   
   //M307EM1
   Z300_Conveyor_Conf[19].dLengthConveyor_cmm := 238000;
   Z300_Conveyor_Conf[19].dWidthConveyor_cmm := 450000;
   Z300_Conveyor_Conf[19].dPitchRoller := 25000;
   Z300_Conveyor_Conf[19].dSpaceRestartPlate_cmm := 200000;
   Z300_Conveyor_Conf[19].dMachineIndex := 19;
   Z300_Conveyor_Conf[19].dZoneConveyor := 1; //Z301
   Z300_Conveyor_Conf[19].dMotorNumber := 0; //Single motor
   Z300_Conveyor_Conf[19].dIndexMainSpeed := 0; //Auto speed
   Z300_Conveyor_Conf[19].xContinuousConveyor := 0;
   Z300_Conveyor_Conf[19].xWaitGlassForStop := 1;
   Z300_Conveyor_Conf[19].rAccH_ms2 := 1.2;
   Z300_Conveyor_Conf[19].rDecH_ms2 := 1.2;
   Z300_Conveyor_Conf[19].rAccH_s := 1.25; //acceleration time with max speed 90 m/min
   Z300_Conveyor_Conf[19].rDecH_s := 1.25; //acceleration time with max speed 90 m/min
   Z300_Conveyor_Conf[19].rAccL_ms2 := 0.7;
   Z300_Conveyor_Conf[19].rDecL_ms2 := 0.7;
   Z300_Conveyor_Conf[19].rAccL_s := 2.14; //acceleration time with max speed 90 m/min
   Z300_Conveyor_Conf[19].rDecL_s := 2.14; //acceleration time with max speed 90 m/min
   Z300_Conveyor_Conf[19].xSimulationMotor := TMP_xSimulationActive;
   Z300_Conveyor_Conf[19].xLocalCleaningAllow := 0;
   Z300_Conveyor_Conf[19].xOnlyOnePlateAtTheTime := 0;
   Z300_Conveyor_Conf[19].rgxAllowedDest := CONST_rgdDestMask[0] AND CONST_rgdDestMask[1] AND CONST_rgdDestMask[2] AND CONST_rgdDestMask[3] AND CONST_rgdDestMask[4] AND CONST_rgdDestMask[5] AND CONST_rgdDestMask[6];
   Z300_Conveyor_Conf[19].rgxAllowedCullet := CONST_rgdDestMask[24];
   Z300_Conveyor_Conf[19].rgxAllowedQuality := CONST_rgdDestMask[29] AND CONST_rgdDestMask[30] AND CONST_rgdDestMask[31];
   Z300_Conveyor[19].tmOFF_DriveEnable[0].PRE := 30000;
   Z300_Conveyor[19].tmON_FeedbackTimeout[0].PRE := 2500;
   Z300_Conveyor[19].tmON_FeedbackTimeout[1].PRE := 2500;
   Z300_Conveyor[19].tmON_DelayReadyToMove[0].PRE := 200;
   Z300_Conveyor[19].tmON_DelayReadyToMove[1].PRE := 200;
   Z300_Conveyor[19].tmON_FeedbackDriveReady[0].PRE := 1000;
   Z300_Conveyor[19].tmON_FeedbackDriveReady[1].PRE := 1000;
   
   //M307FM1
   Z300_Conveyor_Conf[20].dLengthConveyor_cmm := 238000;
   Z300_Conveyor_Conf[20].dWidthConveyor_cmm := 450000;
   Z300_Conveyor_Conf[20].dPitchRoller := 25000;
   Z300_Conveyor_Conf[20].dSpaceRestartPlate_cmm := 200000;
   Z300_Conveyor_Conf[20].dMachineIndex := 20;
   Z300_Conveyor_Conf[20].dZoneConveyor := 1; //Z301
   Z300_Conveyor_Conf[20].dMotorNumber := 0; //Single motor
   Z300_Conveyor_Conf[20].dIndexMainSpeed := 0; //Auto speed
   Z300_Conveyor_Conf[20].xContinuousConveyor := 0;
   Z300_Conveyor_Conf[20].xWaitGlassForStop := 1;
   Z300_Conveyor_Conf[20].rAccH_ms2 := 1.2;
   Z300_Conveyor_Conf[20].rDecH_ms2 := 1.2;
   Z300_Conveyor_Conf[20].rAccH_s := 1.25; //acceleration time with max speed 90 m/min
   Z300_Conveyor_Conf[20].rDecH_s := 1.25; //acceleration time with max speed 90 m/min
   Z300_Conveyor_Conf[20].rAccL_ms2 := 0.7;
   Z300_Conveyor_Conf[20].rDecL_ms2 := 0.7;
   Z300_Conveyor_Conf[20].rAccL_s := 2.14; //acceleration time with max speed 90 m/min
   Z300_Conveyor_Conf[20].rDecL_s := 2.14; //acceleration time with max speed 90 m/min
   Z300_Conveyor_Conf[20].xSimulationMotor := TMP_xSimulationActive;
   Z300_Conveyor_Conf[20].xLocalCleaningAllow := 0;
   Z300_Conveyor_Conf[20].xOnlyOnePlateAtTheTime := 0;
   Z300_Conveyor_Conf[20].rgxAllowedDest := CONST_rgdDestMask[0] AND CONST_rgdDestMask[1] AND CONST_rgdDestMask[2] AND CONST_rgdDestMask[3] AND CONST_rgdDestMask[4] AND CONST_rgdDestMask[5] AND CONST_rgdDestMask[6];
   Z300_Conveyor_Conf[20].rgxAllowedCullet := CONST_rgdDestMask[24];
   Z300_Conveyor_Conf[20].rgxAllowedQuality := CONST_rgdDestMask[29] AND CONST_rgdDestMask[30] AND CONST_rgdDestMask[31];
   Z300_Conveyor[20].tmOFF_DriveEnable[0].PRE := 30000;
   Z300_Conveyor[20].tmON_FeedbackTimeout[0].PRE := 2500;
   Z300_Conveyor[20].tmON_DelayReadyToMove[0].PRE := 200;
   Z300_Conveyor[20].tmON_FeedbackDriveReady[0].PRE := 1000;
   
   //M350M1
   Z300_Conveyor_Conf[21].dLengthConveyor_cmm := 237000;
   Z300_Conveyor_Conf[21].dWidthConveyor_cmm := 450000;
   Z300_Conveyor_Conf[21].dPitchRoller := 25000;
   Z300_Conveyor_Conf[21].dSpaceRestartPlate_cmm := 200000;
   Z300_Conveyor_Conf[21].dMachineIndex := 21;
   Z300_Conveyor_Conf[21].dZoneConveyor := 1; //Z301
   Z300_Conveyor_Conf[21].dMotorNumber := 0; //Single motor
   Z300_Conveyor_Conf[21].dIndexMainSpeed := 0; //Auto speed
   Z300_Conveyor_Conf[21].xContinuousConveyor := 0;
   Z300_Conveyor_Conf[21].xWaitGlassForStop := 1;
   Z300_Conveyor_Conf[21].rAccH_ms2 := 1.2;
   Z300_Conveyor_Conf[21].rDecH_ms2 := 1.2;
   Z300_Conveyor_Conf[21].rAccH_s := 1.25; //acceleration time with max speed 90 m/min
   Z300_Conveyor_Conf[21].rDecH_s := 1.25; //acceleration time with max speed 90 m/min
   Z300_Conveyor_Conf[21].rAccL_ms2 := 0.7;
   Z300_Conveyor_Conf[21].rDecL_ms2 := 0.7;
   Z300_Conveyor_Conf[21].rAccL_s := 2.14; //acceleration time with max speed 90 m/min
   Z300_Conveyor_Conf[21].rDecL_s := 2.14; //acceleration time with max speed 90 m/min
   Z300_Conveyor_Conf[21].xSimulationMotor := TMP_xSimulationActive;
   Z300_Conveyor_Conf[21].xLocalCleaningAllow := 0;
   Z300_Conveyor_Conf[21].xOnlyOnePlateAtTheTime := 0;
   Z300_Conveyor_Conf[21].rgxAllowedDest := CONST_rgdDestMask[0] AND CONST_rgdDestMask[1] AND CONST_rgdDestMask[2] AND CONST_rgdDestMask[3] AND CONST_rgdDestMask[4] AND CONST_rgdDestMask[5] AND CONST_rgdDestMask[6];
   Z300_Conveyor_Conf[21].rgxAllowedCullet := CONST_rgdDestMask[24];
   Z300_Conveyor_Conf[21].rgxAllowedQuality := CONST_rgdDestMask[29] AND CONST_rgdDestMask[30] AND CONST_rgdDestMask[31];
   Z300_Conveyor[21].tmOFF_DriveEnable[0].PRE := 30000;
   Z300_Conveyor[21].tmON_FeedbackTimeout[0].PRE := 2500;
   Z300_Conveyor[21].tmON_DelayReadyToMove[0].PRE := 200;
   Z300_Conveyor[21].tmON_FeedbackDriveReady[0].PRE := 1000;
   
   //M310M1
   Z300_Conveyor_Conf[22].dLengthConveyor_cmm := 243000;
   Z300_Conveyor_Conf[22].dWidthConveyor_cmm := 450000;
   Z300_Conveyor_Conf[22].dPitchRoller := 25000;
   Z300_Conveyor_Conf[22].dSpaceRestartPlate_cmm := 200000;
   Z300_Conveyor_Conf[22].dMachineIndex := 22;
   Z300_Conveyor_Conf[22].dZoneConveyor := 1; //Z301
   Z300_Conveyor_Conf[22].dMotorNumber := 0; //Single motor
   Z300_Conveyor_Conf[22].dIndexMainSpeed := 0; //Auto speed
   Z300_Conveyor_Conf[22].xContinuousConveyor := 0;
   Z300_Conveyor_Conf[22].xWaitGlassForStop := 1;
   Z300_Conveyor_Conf[22].rAccH_ms2 := 1.2;
   Z300_Conveyor_Conf[22].rDecH_ms2 := 1.2;
   Z300_Conveyor_Conf[22].rAccH_s := 1.25; //acceleration time with max speed 90 m/min
   Z300_Conveyor_Conf[22].rDecH_s := 1.25; //acceleration time with max speed 90 m/min
   Z300_Conveyor_Conf[22].rAccL_ms2 := 0.7;
   Z300_Conveyor_Conf[22].rDecL_ms2 := 0.7;
   Z300_Conveyor_Conf[22].rAccL_s := 2.14; //acceleration time with max speed 90 m/min
   Z300_Conveyor_Conf[22].rDecL_s := 2.14; //acceleration time with max speed 90 m/min
   Z300_Conveyor_Conf[22].xSimulationMotor := TMP_xSimulationActive;
   Z300_Conveyor_Conf[22].xLocalCleaningAllow := 0;
   Z300_Conveyor_Conf[22].xOnlyOnePlateAtTheTime := 0;
   Z300_Conveyor_Conf[22].rgxAllowedDest := CONST_rgdDestMask[0] AND CONST_rgdDestMask[1] AND CONST_rgdDestMask[2] AND CONST_rgdDestMask[3] AND CONST_rgdDestMask[4] AND CONST_rgdDestMask[5] AND CONST_rgdDestMask[6];
   Z300_Conveyor_Conf[22].rgxAllowedCullet := CONST_rgdDestMask[24];
   Z300_Conveyor_Conf[22].rgxAllowedQuality := CONST_rgdDestMask[31];
   Z300_Conveyor[22].tmOFF_DriveEnable[0].PRE := 30000;
   Z300_Conveyor[22].tmON_FeedbackTimeout[0].PRE := 2500;
   Z300_Conveyor[22].tmON_DelayReadyToMove[0].PRE := 200;
   Z300_Conveyor[22].tmON_FeedbackDriveReady[0].PRE := 1000;
   
   //M310M2
   Z300_Conveyor_Conf[23].dLengthConveyor_cmm := 243000;
   Z300_Conveyor_Conf[23].dWidthConveyor_cmm := 450000;
   Z300_Conveyor_Conf[23].dPitchRoller := 25000;
   Z300_Conveyor_Conf[23].dSpaceRestartPlate_cmm := 200000;
   Z300_Conveyor_Conf[23].dMachineIndex := 23;
   Z300_Conveyor_Conf[23].dZoneConveyor := 1; //Z301
   Z300_Conveyor_Conf[23].dMotorNumber := 0; //Single motor
   Z300_Conveyor_Conf[23].dIndexMainSpeed := 0; //Auto speed
   Z300_Conveyor_Conf[23].xContinuousConveyor := 0;
   Z300_Conveyor_Conf[23].xWaitGlassForStop := 1;
   Z300_Conveyor_Conf[23].rAccH_ms2 := 1.2;
   Z300_Conveyor_Conf[23].rDecH_ms2 := 1.2;
   Z300_Conveyor_Conf[23].rAccH_s := 1.25; //acceleration time with max speed 90 m/min
   Z300_Conveyor_Conf[23].rDecH_s := 1.25; //acceleration time with max speed 90 m/min
   Z300_Conveyor_Conf[23].rAccL_ms2 := 0.7;
   Z300_Conveyor_Conf[23].rDecL_ms2 := 0.7;
   Z300_Conveyor_Conf[23].rAccL_s := 2.14; //acceleration time with max speed 90 m/min
   Z300_Conveyor_Conf[23].rDecL_s := 2.14; //acceleration time with max speed 90 m/min
   Z300_Conveyor_Conf[23].xSimulationMotor := TMP_xSimulationActive;
   Z300_Conveyor_Conf[23].xLocalCleaningAllow := 0;
   Z300_Conveyor_Conf[23].xOnlyOnePlateAtTheTime := 0;
   Z300_Conveyor_Conf[23].rgxAllowedDest := CONST_rgdDestMask[0] AND CONST_rgdDestMask[1] AND CONST_rgdDestMask[2] AND CONST_rgdDestMask[3] AND CONST_rgdDestMask[4] AND CONST_rgdDestMask[5] AND CONST_rgdDestMask[6];
   Z300_Conveyor_Conf[23].rgxAllowedCullet := CONST_rgdDestMask[24];
   Z300_Conveyor_Conf[23].rgxAllowedQuality := CONST_rgdDestMask[31];
   Z300_Conveyor[23].tmOFF_DriveEnable[0].PRE := 30000;
   Z300_Conveyor[23].tmON_FeedbackTimeout[0].PRE := 2500;
   Z300_Conveyor[23].tmON_DelayReadyToMove[0].PRE := 200;
   Z300_Conveyor[23].tmON_FeedbackDriveReady[0].PRE := 1000;
   
   //M310M3
   Z300_Conveyor_Conf[24].dLengthConveyor_cmm := 243000;
   Z300_Conveyor_Conf[24].dWidthConveyor_cmm := 450000;
   Z300_Conveyor_Conf[24].dPitchRoller := 25000;
   Z300_Conveyor_Conf[24].dSpaceRestartPlate_cmm := 200000;
   Z300_Conveyor_Conf[24].dMachineIndex := 24;
   Z300_Conveyor_Conf[24].dZoneConveyor := 1; //Z301
   Z300_Conveyor_Conf[24].dMotorNumber := 0; //Single motor
   Z300_Conveyor_Conf[24].dIndexMainSpeed := 0; //Auto speed
   Z300_Conveyor_Conf[24].xContinuousConveyor := 0;
   Z300_Conveyor_Conf[24].xWaitGlassForStop := 1;
   Z300_Conveyor_Conf[24].rAccH_ms2 := 1.2;
   Z300_Conveyor_Conf[24].rDecH_ms2 := 1.2;
   Z300_Conveyor_Conf[24].rAccH_s := 1.25; //acceleration time with max speed 90 m/min
   Z300_Conveyor_Conf[24].rDecH_s := 1.25; //acceleration time with max speed 90 m/min
   Z300_Conveyor_Conf[24].rAccL_ms2 := 0.7;
   Z300_Conveyor_Conf[24].rDecL_ms2 := 0.7;
   Z300_Conveyor_Conf[24].rAccL_s := 2.14; //acceleration time with max speed 90 m/min
   Z300_Conveyor_Conf[24].rDecL_s := 2.14; //acceleration time with max speed 90 m/min
   Z300_Conveyor_Conf[24].xSimulationMotor := TMP_xSimulationActive;
   Z300_Conveyor_Conf[24].xLocalCleaningAllow := 0;
   Z300_Conveyor_Conf[24].xOnlyOnePlateAtTheTime := 0;
   Z300_Conveyor_Conf[24].rgxAllowedDest := CONST_rgdDestMask[0] AND CONST_rgdDestMask[1] AND CONST_rgdDestMask[2] AND CONST_rgdDestMask[3] AND CONST_rgdDestMask[4] AND CONST_rgdDestMask[5] AND CONST_rgdDestMask[6];
   Z300_Conveyor_Conf[24].rgxAllowedCullet := CONST_rgdDestMask[24];
   Z300_Conveyor_Conf[24].rgxAllowedQuality := CONST_rgdDestMask[31];
   Z300_Conveyor[24].tmOFF_DriveEnable[0].PRE := 30000;
   Z300_Conveyor[24].tmON_FeedbackTimeout[0].PRE := 2500;
   Z300_Conveyor[24].tmON_DelayReadyToMove[0].PRE := 200;
   Z300_Conveyor[24].tmON_FeedbackDriveReady[0].PRE := 1000;
   
   //M360M1
   Z300_Conveyor_Conf[25].dLengthConveyor_cmm := 393000;
   Z300_Conveyor_Conf[25].dWidthConveyor_cmm := 450000;
   Z300_Conveyor_Conf[25].dPitchRoller := 25000;
   Z300_Conveyor_Conf[25].dSpaceRestartPlate_cmm := 350000;
   Z300_Conveyor_Conf[25].dMachineIndex := 25;
   Z300_Conveyor_Conf[25].dZoneConveyor := 1; //Z301
   Z300_Conveyor_Conf[25].dMotorNumber := 0; //Single motor
   Z300_Conveyor_Conf[25].dIndexMainSpeed := 0; //Auto speed
   Z300_Conveyor_Conf[25].xContinuousConveyor := 0;
   Z300_Conveyor_Conf[25].xWaitGlassForStop := 1;
   Z300_Conveyor_Conf[25].rAccH_ms2 := 1.2;
   Z300_Conveyor_Conf[25].rDecH_ms2 := 1.2;
   Z300_Conveyor_Conf[25].rAccH_s := 1.25; //acceleration time with max speed 90 m/min
   Z300_Conveyor_Conf[25].rDecH_s := 1.25; //acceleration time with max speed 90 m/min
   Z300_Conveyor_Conf[25].rAccL_ms2 := 0.7;
   Z300_Conveyor_Conf[25].rDecL_ms2 := 0.7;
   Z300_Conveyor_Conf[25].rAccL_s := 2.14; //acceleration time with max speed 90 m/min
   Z300_Conveyor_Conf[25].rDecL_s := 2.14; //acceleration time with max speed 90 m/min
   Z300_Conveyor_Conf[25].xSimulationMotor := TMP_xSimulationActive;
   Z300_Conveyor_Conf[25].xLocalCleaningAllow := 0;
   Z300_Conveyor_Conf[25].xOnlyOnePlateAtTheTime := 0;
   Z300_Conveyor_Conf[25].rgxAllowedDest := CONST_rgdDestMask[1] AND CONST_rgdDestMask[2] AND CONST_rgdDestMask[3] AND CONST_rgdDestMask[4] AND CONST_rgdDestMask[5] AND CONST_rgdDestMask[6];
   Z300_Conveyor_Conf[25].rgxAllowedCullet := CONST_rgdDestMask[24];
   Z300_Conveyor_Conf[25].rgxAllowedQuality := CONST_rgdDestMask[31];
   Z300_Conveyor[25].tmOFF_DriveEnable[0].PRE := 30000;
   Z300_Conveyor[25].tmON_FeedbackTimeout[0].PRE := 2500;
   Z300_Conveyor[25].tmON_DelayReadyToMove[0].PRE := 200;
   Z300_Conveyor[25].tmON_FeedbackDriveReady[0].PRE := 1000;
   
   //M315M1
   Z300_Conveyor_Conf[26].dLengthConveyor_cmm := 243000;
   Z300_Conveyor_Conf[26].dWidthConveyor_cmm := 450000;
   Z300_Conveyor_Conf[26].dPitchRoller := 25000;
   Z300_Conveyor_Conf[26].dSpaceRestartPlate_cmm := 200000;
   Z300_Conveyor_Conf[26].dMachineIndex := 26;
   Z300_Conveyor_Conf[26].dZoneConveyor := 1; //Z301
   Z300_Conveyor_Conf[26].dMotorNumber := 0; //Single motor
   Z300_Conveyor_Conf[26].dIndexMainSpeed := 0; //Auto speed
   Z300_Conveyor_Conf[26].xContinuousConveyor := 0;
   Z300_Conveyor_Conf[26].xWaitGlassForStop := 1;
   Z300_Conveyor_Conf[26].rAccH_ms2 := 1.2;
   Z300_Conveyor_Conf[26].rDecH_ms2 := 1.2;
   Z300_Conveyor_Conf[26].rAccH_s := 1.25; //acceleration time with max speed 90 m/min
   Z300_Conveyor_Conf[26].rDecH_s := 1.25; //acceleration time with max speed 90 m/min
   Z300_Conveyor_Conf[26].rAccL_ms2 := 0.7;
   Z300_Conveyor_Conf[26].rDecL_ms2 := 0.7;
   Z300_Conveyor_Conf[26].rAccL_s := 2.14; //acceleration time with max speed 90 m/min
   Z300_Conveyor_Conf[26].rDecL_s := 2.14; //acceleration time with max speed 90 m/min
   Z300_Conveyor_Conf[26].xSimulationMotor := TMP_xSimulationActive;
   Z300_Conveyor_Conf[26].xLocalCleaningAllow := 0;
   Z300_Conveyor_Conf[26].xOnlyOnePlateAtTheTime := 0;
   Z300_Conveyor_Conf[26].rgxAllowedDest := CONST_rgdDestMask[1] AND CONST_rgdDestMask[2] AND CONST_rgdDestMask[3] AND CONST_rgdDestMask[4] AND CONST_rgdDestMask[5] AND CONST_rgdDestMask[6];
   Z300_Conveyor_Conf[26].rgxAllowedCullet := CONST_rgdDestMask[24];
   Z300_Conveyor_Conf[26].rgxAllowedQuality := CONST_rgdDestMask[31];
   Z300_Conveyor[26].tmOFF_DriveEnable[0].PRE := 30000;
   Z300_Conveyor[26].tmON_FeedbackTimeout[0].PRE := 2500;
   Z300_Conveyor[26].tmON_DelayReadyToMove[0].PRE := 200;
   Z300_Conveyor[26].tmON_FeedbackDriveReady[0].PRE := 1000;
   
   //M315M2
   Z300_Conveyor_Conf[27].dLengthConveyor_cmm := 243000;
   Z300_Conveyor_Conf[27].dWidthConveyor_cmm := 450000;
   Z300_Conveyor_Conf[27].dPitchRoller := 25000;
   Z300_Conveyor_Conf[27].dSpaceRestartPlate_cmm := 200000;
   Z300_Conveyor_Conf[27].dMachineIndex := 27;
   Z300_Conveyor_Conf[27].dZoneConveyor := 1; //Z301
   Z300_Conveyor_Conf[27].dMotorNumber := 0; //Single motor
   Z300_Conveyor_Conf[27].dIndexMainSpeed := 0; //Auto speed
   Z300_Conveyor_Conf[27].xContinuousConveyor := 1;
   Z300_Conveyor_Conf[27].xWaitGlassForStop := 1;
   Z300_Conveyor_Conf[27].rAccH_ms2 := 1.2;
   Z300_Conveyor_Conf[27].rDecH_ms2 := 1.2;
   Z300_Conveyor_Conf[27].rAccH_s := 1.25; //acceleration time with max speed 90 m/min
   Z300_Conveyor_Conf[27].rDecH_s := 1.25; //acceleration time with max speed 90 m/min
   Z300_Conveyor_Conf[27].rAccL_ms2 := 0.7;
   Z300_Conveyor_Conf[27].rDecL_ms2 := 0.7;
   Z300_Conveyor_Conf[27].rAccL_s := 2.14; //acceleration time with max speed 90 m/min
   Z300_Conveyor_Conf[27].rDecL_s := 2.14; //acceleration time with max speed 90 m/min
   Z300_Conveyor_Conf[27].xSimulationMotor := TMP_xSimulationActive;
   Z300_Conveyor_Conf[27].xLocalCleaningAllow := 0;
   Z300_Conveyor_Conf[27].xOnlyOnePlateAtTheTime := 0;
   Z300_Conveyor_Conf[27].rgxAllowedDest := CONST_rgdDestMask[1] AND CONST_rgdDestMask[2] AND CONST_rgdDestMask[3] AND CONST_rgdDestMask[4] AND CONST_rgdDestMask[5] AND CONST_rgdDestMask[6];
   Z300_Conveyor_Conf[27].rgxAllowedCullet := CONST_rgdDestMask[24];
   Z300_Conveyor_Conf[27].rgxAllowedQuality := CONST_rgdDestMask[31];
   Z300_Conveyor[27].tmOFF_DriveEnable[0].PRE := 30000;
   Z300_Conveyor[27].tmON_FeedbackTimeout[0].PRE := 2500;
   Z300_Conveyor[27].tmON_DelayReadyToMove[0].PRE := 200;
   Z300_Conveyor[27].tmON_FeedbackDriveReady[0].PRE := 1000;
   
   //M315M3
   Z300_Conveyor_Conf[28].dLengthConveyor_cmm := 243000;
   Z300_Conveyor_Conf[28].dWidthConveyor_cmm := 450000;
   Z300_Conveyor_Conf[28].dPitchRoller := 25000;
   Z300_Conveyor_Conf[28].dSpaceRestartPlate_cmm := 200000;
   Z300_Conveyor_Conf[28].dMachineIndex := 28;
   Z300_Conveyor_Conf[28].dZoneConveyor := 1; //Z301
   Z300_Conveyor_Conf[28].dMotorNumber := 0; //Single motor
   Z300_Conveyor_Conf[28].dIndexMainSpeed := 0; //Auto speed
   Z300_Conveyor_Conf[28].xContinuousConveyor := 1;
   Z300_Conveyor_Conf[28].xWaitGlassForStop := 1;
   Z300_Conveyor_Conf[28].rAccH_ms2 := 1.2;
   Z300_Conveyor_Conf[28].rDecH_ms2 := 1.2;
   Z300_Conveyor_Conf[28].rAccH_s := 1.25; //acceleration time with max speed 90 m/min
   Z300_Conveyor_Conf[28].rDecH_s := 1.25; //acceleration time with max speed 90 m/min
   Z300_Conveyor_Conf[28].rAccL_ms2 := 0.7;
   Z300_Conveyor_Conf[28].rDecL_ms2 := 0.7;
   Z300_Conveyor_Conf[28].rAccL_s := 2.14; //acceleration time with max speed 90 m/min
   Z300_Conveyor_Conf[28].rDecL_s := 2.14; //acceleration time with max speed 90 m/min
   Z300_Conveyor_Conf[28].xSimulationMotor := TMP_xSimulationActive;
   Z300_Conveyor_Conf[28].xLocalCleaningAllow := 0;
   Z300_Conveyor_Conf[28].xOnlyOnePlateAtTheTime := 0;
   Z300_Conveyor_Conf[28].rgxAllowedDest := CONST_rgdDestMask[1] AND CONST_rgdDestMask[2] AND CONST_rgdDestMask[3] AND CONST_rgdDestMask[4] AND CONST_rgdDestMask[5] AND CONST_rgdDestMask[6];
   Z300_Conveyor_Conf[28].rgxAllowedCullet := CONST_rgdDestMask[24];
   Z300_Conveyor_Conf[28].rgxAllowedQuality := CONST_rgdDestMask[31];
   Z300_Conveyor[28].tmOFF_DriveEnable[0].PRE := 30000;
   Z300_Conveyor[28].tmON_FeedbackTimeout[0].PRE := 2500;
   Z300_Conveyor[28].tmON_DelayReadyToMove[0].PRE := 200;
   Z300_Conveyor[28].tmON_FeedbackDriveReady[0].PRE := 1000;
   
   
END_ROUTINE

ROUTINE Conv_Faults   (* ladder *)
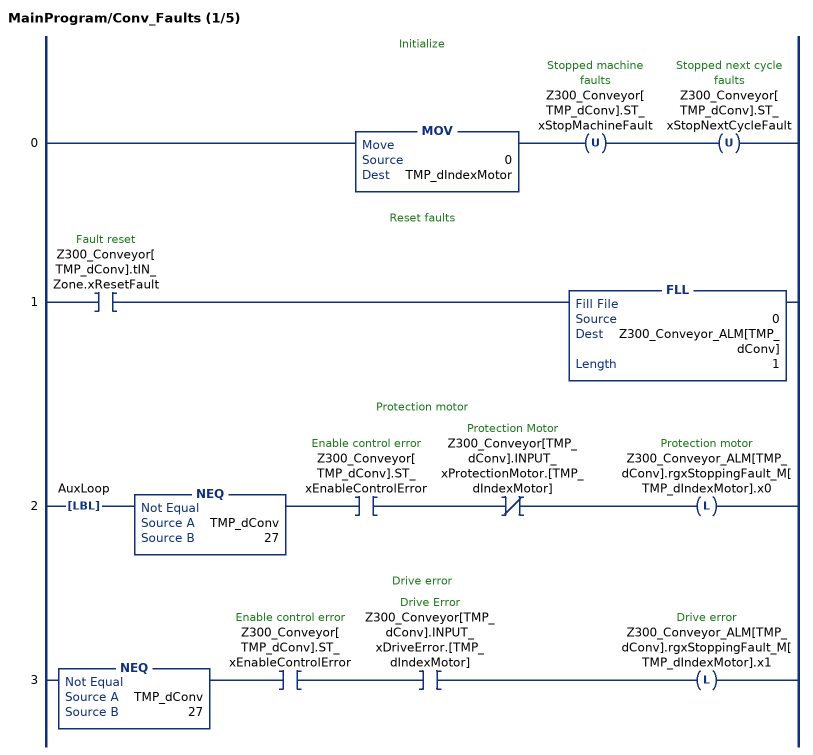
   // Initialize
   0: MOV(0,TMP_dIndexMotor)OTU(Z300_Conveyor[TMP_dConv].ST_xStopMachineFault)OTU(Z300_Conveyor[TMP_dConv].ST_xStopNextCycleFault);
   // Reset faults
   1: XIC(Z300_Conveyor[TMP_dConv].tIN_Zone.xResetFault)FLL(0,Z300_Conveyor_ALM[TMP_dConv],1);
   // Protection motor
   2: LBL(AuxLoop)NEQ(TMP_dConv,27)XIC(Z300_Conveyor[TMP_dConv].ST_xEnableControlError)XIO(Z300_Conveyor[TMP_dConv].INPUT_xProtectionMotor.[TMP_dIndexMotor])OTL(Z300_Conveyor_ALM[TMP_dConv].rgxStoppingFault_M[TMP_dIndexMotor].x0);
   // Drive error
   3: NEQ(TMP_dConv,27)XIC(Z300_Conveyor[TMP_dConv].ST_xEnableControlError)XIC(Z300_Conveyor[TMP_dConv].INPUT_xDriveError.[TMP_dIndexMotor])OTL(Z300_Conveyor_ALM[TMP_dConv].rgxStoppingFault_M[TMP_dIndexMotor].x1);
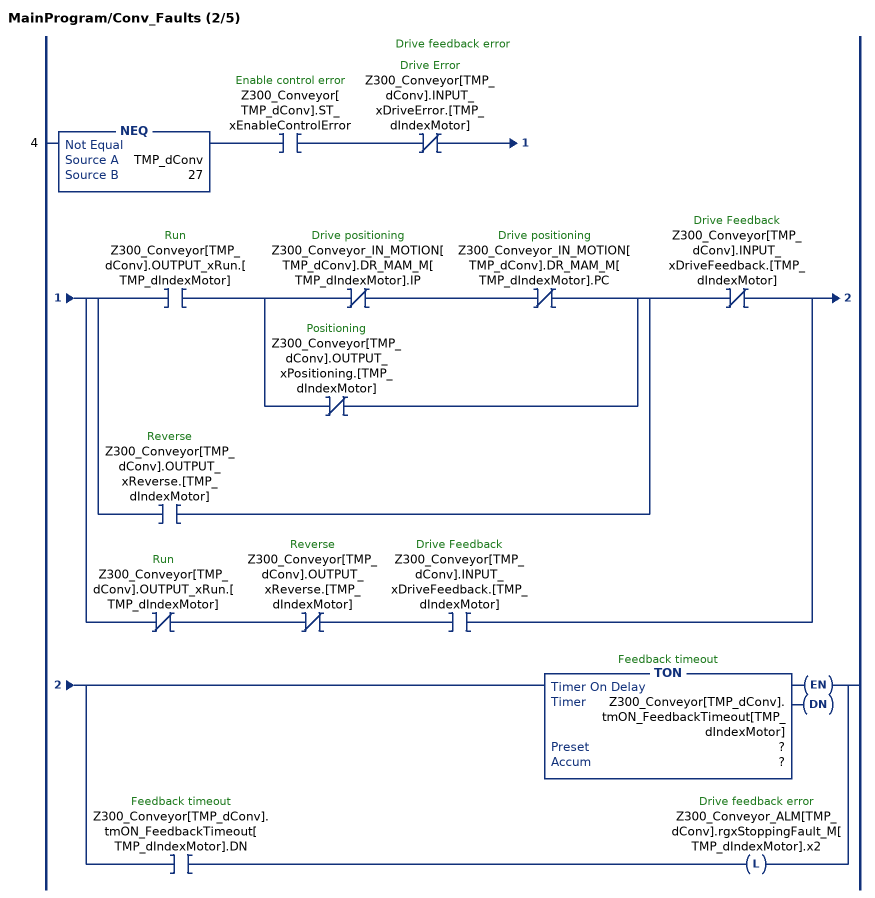
   // Drive feedback error
   4: NEQ(TMP_dConv,27)XIC(Z300_Conveyor[TMP_dConv].ST_xEnableControlError)XIO(Z300_Conveyor[TMP_dConv].INPUT_xDriveError.[TMP_dIndexMotor])[[XIC(Z300_Conveyor[TMP_dConv].OUTPUT_xRun.[TMP_dIndexMotor]) [XIO(Z300_Conveyor_IN_MOTION[TMP_dConv].DR_MAM_M[TMP_dIndexMotor].IP) XIO(Z300_Conveyor_IN_MOTION[TMP_dConv].DR_MAM_M[TMP_dIndexMotor].PC) ,XIO(Z300_Conveyor[TMP_dConv].OUTPUT_xPositioning.[TMP_dIndexMotor]) ] ,XIC(Z300_Conveyor[TMP_dConv].OUTPUT_xReverse.[TMP_dIndexMotor]) ] XIO(Z300_Conveyor[TMP_dConv].INPUT_xDriveFeedback.[TMP_dIndexMotor]) ,XIO(Z300_Conveyor[TMP_dConv].OUTPUT_xRun.[TMP_dIndexMotor]) XIO(Z300_Conveyor[TMP_dConv].OUTPUT_xReverse.[TMP_dIndexMotor]) XIC(Z300_Conveyor[TMP_dConv].INPUT_xDriveFeedback.[TMP_dIndexMotor]) ][TON(Z300_Conveyor[TMP_dConv].tmON_FeedbackTimeout[TMP_dIndexMotor],?,?) ,XIC(Z300_Conveyor[TMP_dConv].tmON_FeedbackTimeout[TMP_dIndexMotor].DN) OTL(Z300_Conveyor_ALM[TMP_dConv].rgxStoppingFault_M[TMP_dIndexMotor].x2) ];
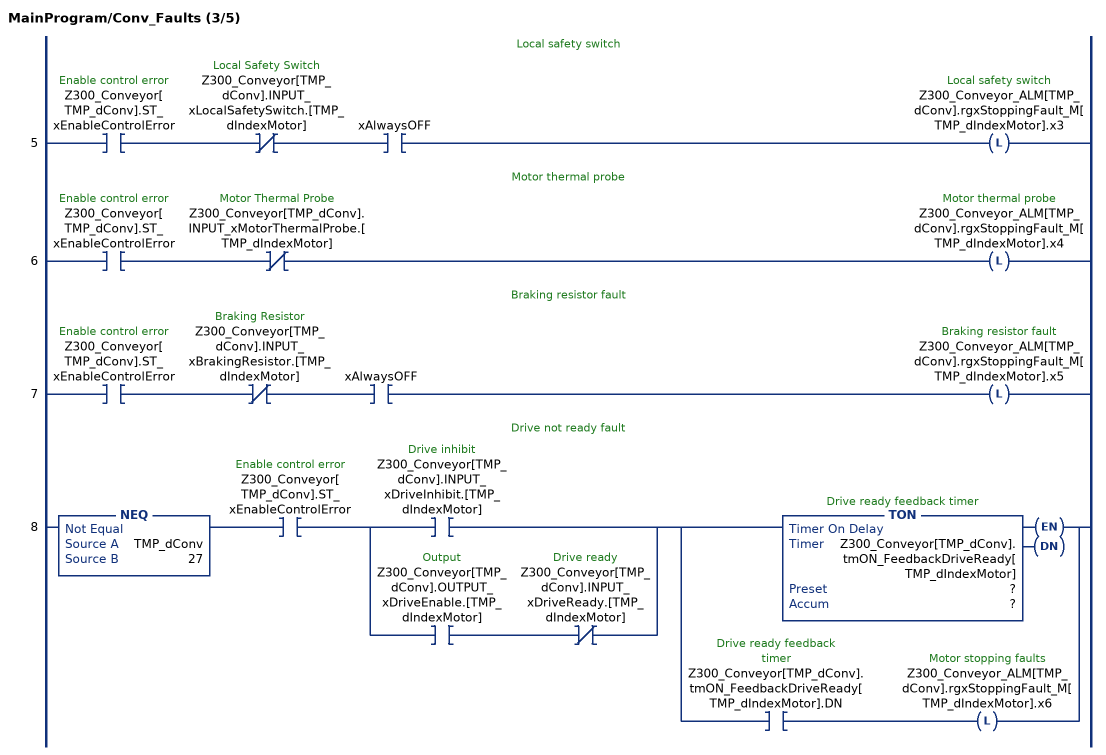
   // Local safety switch
   5: XIC(Z300_Conveyor[TMP_dConv].ST_xEnableControlError)XIO(Z300_Conveyor[TMP_dConv].INPUT_xLocalSafetySwitch.[TMP_dIndexMotor])XIC(xAlwaysOFF)OTL(Z300_Conveyor_ALM[TMP_dConv].rgxStoppingFault_M[TMP_dIndexMotor].x3);
   // Motor thermal probe
   6: XIC(Z300_Conveyor[TMP_dConv].ST_xEnableControlError)XIO(Z300_Conveyor[TMP_dConv].INPUT_xMotorThermalProbe.[TMP_dIndexMotor])OTL(Z300_Conveyor_ALM[TMP_dConv].rgxStoppingFault_M[TMP_dIndexMotor].x4);
   // Braking resistor fault
   7: XIC(Z300_Conveyor[TMP_dConv].ST_xEnableControlError)XIO(Z300_Conveyor[TMP_dConv].INPUT_xBrakingResistor.[TMP_dIndexMotor])XIC(xAlwaysOFF)OTL(Z300_Conveyor_ALM[TMP_dConv].rgxStoppingFault_M[TMP_dIndexMotor].x5);
   // Drive not ready fault
   8: NEQ(TMP_dConv,27)XIC(Z300_Conveyor[TMP_dConv].ST_xEnableControlError)[XIC(Z300_Conveyor[TMP_dConv].INPUT_xDriveInhibit.[TMP_dIndexMotor]) ,XIC(Z300_Conveyor[TMP_dConv].OUTPUT_xDriveEnable.[TMP_dIndexMotor]) XIO(Z300_Conveyor[TMP_dConv].INPUT_xDriveReady.[TMP_dIndexMotor]) ][TON(Z300_Conveyor[TMP_dConv].tmON_FeedbackDriveReady[TMP_dIndexMotor],?,?) ,XIC(Z300_Conveyor[TMP_dConv].tmON_FeedbackDriveReady[TMP_dIndexMotor].DN) OTL(Z300_Conveyor_ALM[TMP_dConv].rgxStoppingFault_M[TMP_dIndexMotor].x6) ];
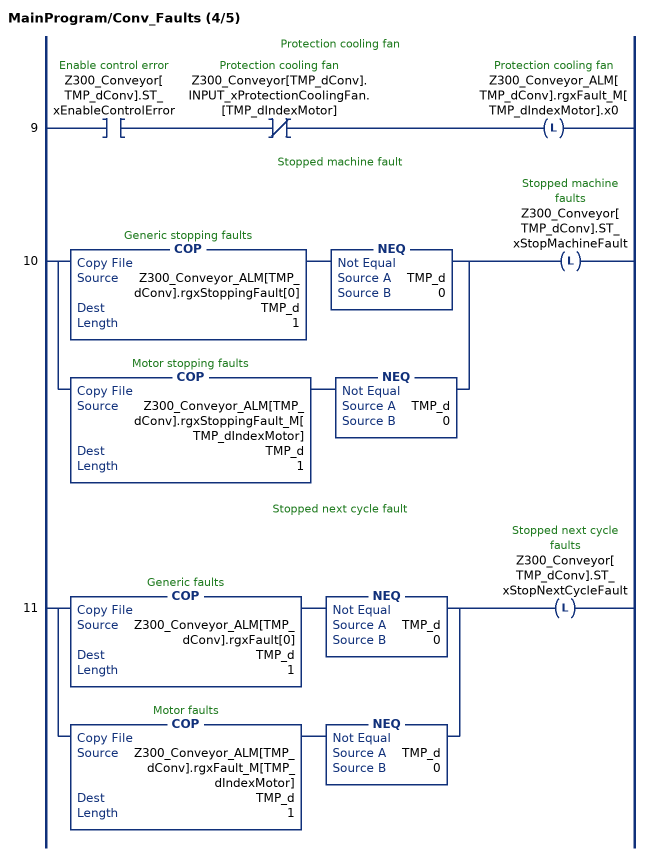
   // Protection cooling fan
   9: XIC(Z300_Conveyor[TMP_dConv].ST_xEnableControlError)XIO(Z300_Conveyor[TMP_dConv].INPUT_xProtectionCoolingFan.[TMP_dIndexMotor])OTL(Z300_Conveyor_ALM[TMP_dConv].rgxFault_M[TMP_dIndexMotor].x0);
   // Stopped machine fault
   10: [COP(Z300_Conveyor_ALM[TMP_dConv].rgxStoppingFault[0],TMP_d,1) NEQ(TMP_d,0) ,COP(Z300_Conveyor_ALM[TMP_dConv].rgxStoppingFault_M[TMP_dIndexMotor],TMP_d,1) NEQ(TMP_d,0) ]OTL(Z300_Conveyor[TMP_dConv].ST_xStopMachineFault);
   // Stopped next cycle fault
   11: [COP(Z300_Conveyor_ALM[TMP_dConv].rgxFault[0],TMP_d,1) NEQ(TMP_d,0) ,COP(Z300_Conveyor_ALM[TMP_dConv].rgxFault_M[TMP_dIndexMotor],TMP_d,1) NEQ(TMP_d,0) ]OTL(Z300_Conveyor[TMP_dConv].ST_xStopNextCycleFault);
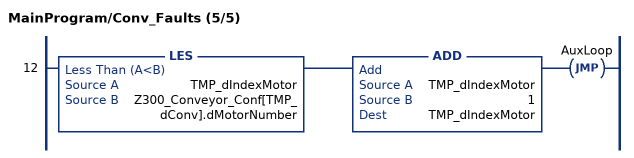
   12: LES(TMP_dIndexMotor,Z300_Conveyor_Conf[TMP_dConv].dMotorNumber)ADD(TMP_dIndexMotor,1,TMP_dIndexMotor)JMP(AuxLoop);
END_ROUTINE

ROUTINE Conv_Logic   (* ladder *)
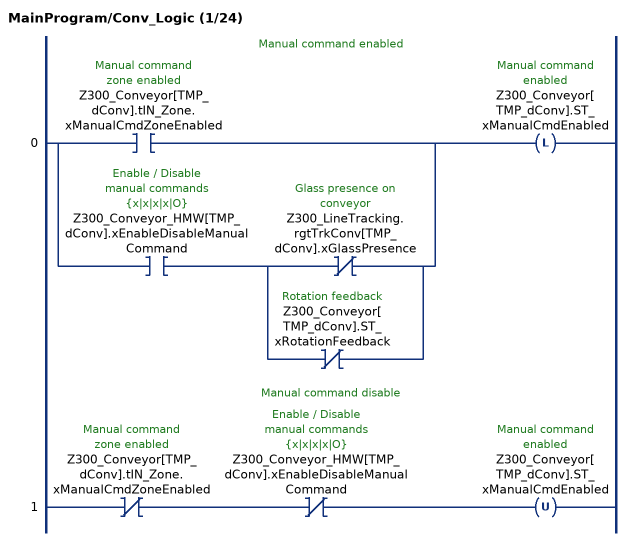
   // Manual command enabled
   0: [XIC(Z300_Conveyor[TMP_dConv].tIN_Zone.xManualCmdZoneEnabled) ,XIC(Z300_Conveyor_HMW[TMP_dConv].xEnableDisableManualCommand) [XIO(Z300_LineTracking.rgtTrkConv[TMP_dConv].xGlassPresence) ,XIO(Z300_Conveyor[TMP_dConv].ST_xRotationFeedback) ] ]OTL(Z300_Conveyor[TMP_dConv].ST_xManualCmdEnabled);
   // Manual command disable
   1: XIO(Z300_Conveyor[TMP_dConv].tIN_Zone.xManualCmdZoneEnabled)XIO(Z300_Conveyor_HMW[TMP_dConv].xEnableDisableManualCommand)OTU(Z300_Conveyor[TMP_dConv].ST_xManualCmdEnabled);
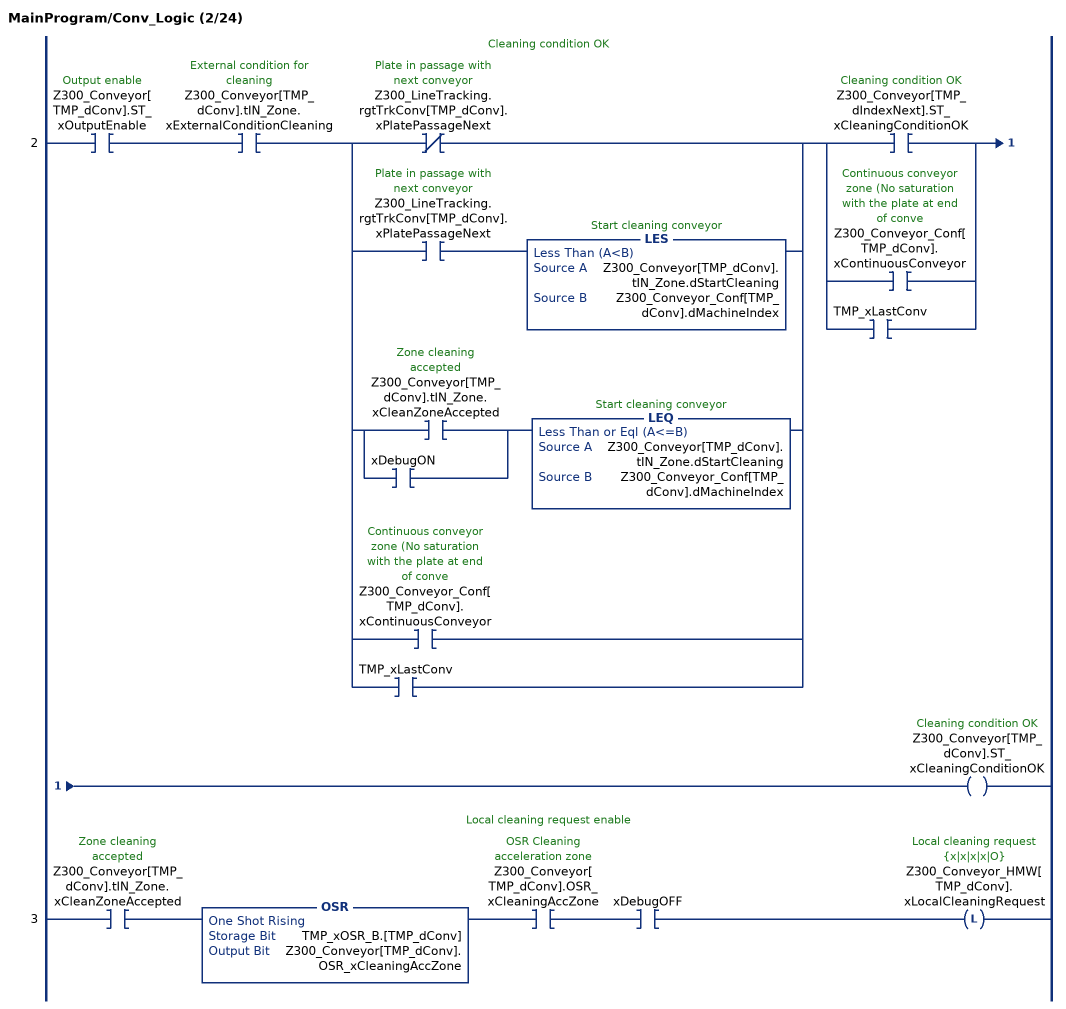
   // Cleaning condition OK
   2: XIC(Z300_Conveyor[TMP_dConv].ST_xOutputEnable)XIC(Z300_Conveyor[TMP_dConv].tIN_Zone.xExternalConditionCleaning)[[XIO(Z300_LineTracking.rgtTrkConv[TMP_dConv].xPlatePassageNext) ,XIC(Z300_LineTracking.rgtTrkConv[TMP_dConv].xPlatePassageNext) LES(Z300_Conveyor[TMP_dConv].tIN_Zone.dStartCleaning,Z300_Conveyor_Conf[TMP_dConv].dMachineIndex) ] ,[[XIC(Z300_Conveyor[TMP_dConv].tIN_Zone.xCleanZoneAccepted) ,XIC(xDebugON) ] LEQ(Z300_Conveyor[TMP_dConv].tIN_Zone.dStartCleaning,Z300_Conveyor_Conf[TMP_dConv].dMachineIndex) ,XIC(Z300_Conveyor_Conf[TMP_dConv].xContinuousConveyor) ,XIC(TMP_xLastConv) ] ][XIC(Z300_Conveyor[TMP_dIndexNext].ST_xCleaningConditionOK) ,[XIC(Z300_Conveyor_Conf[TMP_dConv].xContinuousConveyor) ,XIC(TMP_xLastConv) ] ]OTE(Z300_Conveyor[TMP_dConv].ST_xCleaningConditionOK);
   // Local cleaning request enable
   3: XIC(Z300_Conveyor[TMP_dConv].tIN_Zone.xCleanZoneAccepted)OSR(TMP_xOSR_B.[TMP_dConv],Z300_Conveyor[TMP_dConv].OSR_xCleaningAccZone)XIC(Z300_Conveyor[TMP_dConv].OSR_xCleaningAccZone)XIC(xDebugOFF)OTL(Z300_Conveyor_HMW[TMP_dConv].xLocalCleaningRequest);
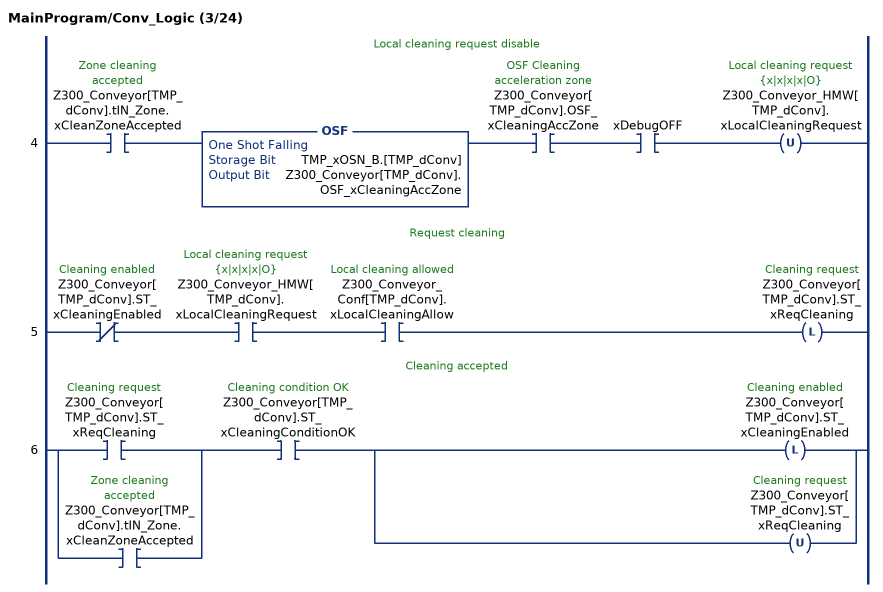
   // Local cleaning request disable
   4: XIC(Z300_Conveyor[TMP_dConv].tIN_Zone.xCleanZoneAccepted)OSF(TMP_xOSN_B.[TMP_dConv],Z300_Conveyor[TMP_dConv].OSF_xCleaningAccZone)XIC(Z300_Conveyor[TMP_dConv].OSF_xCleaningAccZone)XIC(xDebugOFF)OTU(Z300_Conveyor_HMW[TMP_dConv].xLocalCleaningRequest);
   // Request cleaning
   5: XIO(Z300_Conveyor[TMP_dConv].ST_xCleaningEnabled)XIC(Z300_Conveyor_HMW[TMP_dConv].xLocalCleaningRequest)XIC(Z300_Conveyor_Conf[TMP_dConv].xLocalCleaningAllow)OTL(Z300_Conveyor[TMP_dConv].ST_xReqCleaning);
   // Cleaning accepted
   6: [XIC(Z300_Conveyor[TMP_dConv].ST_xReqCleaning) ,XIC(Z300_Conveyor[TMP_dConv].tIN_Zone.xCleanZoneAccepted) ]XIC(Z300_Conveyor[TMP_dConv].ST_xCleaningConditionOK)[OTL(Z300_Conveyor[TMP_dConv].ST_xCleaningEnabled) ,OTU(Z300_Conveyor[TMP_dConv].ST_xReqCleaning) ];
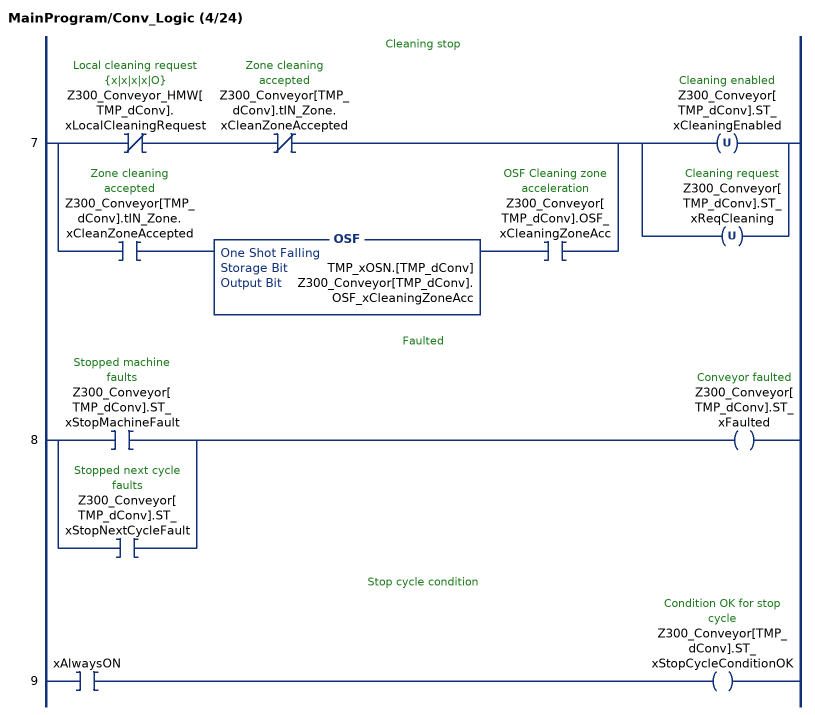
   // Cleaning stop
   7: [XIO(Z300_Conveyor_HMW[TMP_dConv].xLocalCleaningRequest) XIO(Z300_Conveyor[TMP_dConv].tIN_Zone.xCleanZoneAccepted) ,XIC(Z300_Conveyor[TMP_dConv].tIN_Zone.xCleanZoneAccepted) OSF(TMP_xOSN.[TMP_dConv],Z300_Conveyor[TMP_dConv].OSF_xCleaningZoneAcc) XIC(Z300_Conveyor[TMP_dConv].OSF_xCleaningZoneAcc) ][OTU(Z300_Conveyor[TMP_dConv].ST_xCleaningEnabled) ,OTU(Z300_Conveyor[TMP_dConv].ST_xReqCleaning) ];
   // Faulted
   8: [XIC(Z300_Conveyor[TMP_dConv].ST_xStopMachineFault) ,XIC(Z300_Conveyor[TMP_dConv].ST_xStopNextCycleFault) ]OTE(Z300_Conveyor[TMP_dConv].ST_xFaulted);
   // Stop cycle condition
   9: XIC(xAlwaysON)OTE(Z300_Conveyor[TMP_dConv].ST_xStopCycleConditionOK);
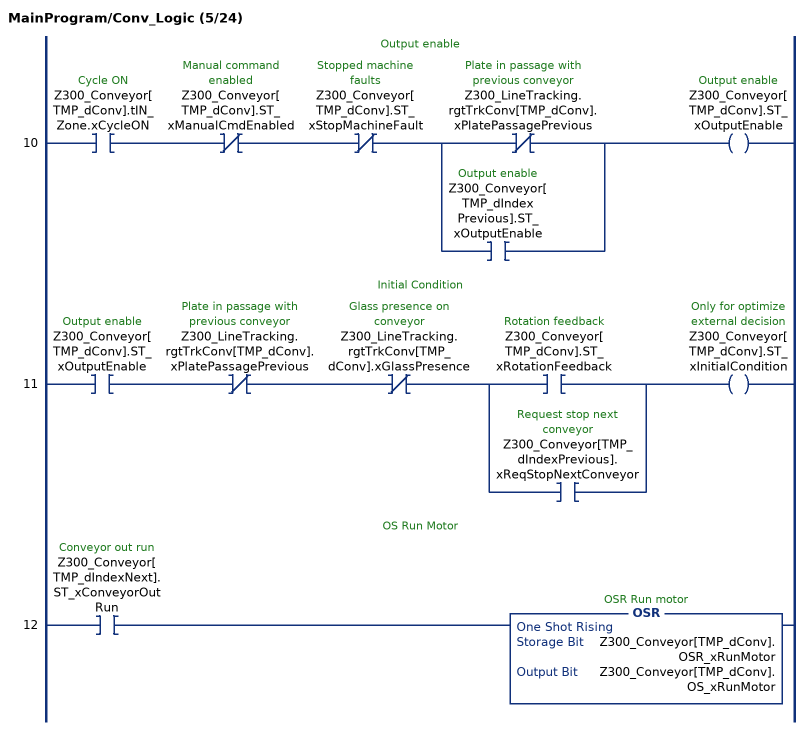
   // Output enable
   10: XIC(Z300_Conveyor[TMP_dConv].tIN_Zone.xCycleON)XIO(Z300_Conveyor[TMP_dConv].ST_xManualCmdEnabled)XIO(Z300_Conveyor[TMP_dConv].ST_xStopMachineFault)[XIO(Z300_LineTracking.rgtTrkConv[TMP_dConv].xPlatePassagePrevious) ,XIC(Z300_Conveyor[TMP_dIndexPrevious].ST_xOutputEnable) ]OTE(Z300_Conveyor[TMP_dConv].ST_xOutputEnable);
   // Initial Condition
   11: XIC(Z300_Conveyor[TMP_dConv].ST_xOutputEnable)XIO(Z300_LineTracking.rgtTrkConv[TMP_dConv].xPlatePassagePrevious)XIO(Z300_LineTracking.rgtTrkConv[TMP_dConv].xGlassPresence)[XIC(Z300_Conveyor[TMP_dConv].ST_xRotationFeedback) ,XIC(Z300_Conveyor[TMP_dIndexPrevious].xReqStopNextConveyor) ]OTE(Z300_Conveyor[TMP_dConv].ST_xInitialCondition);
   // OS Run Motor
   12: XIC(Z300_Conveyor[TMP_dIndexNext].ST_xConveyorOutRun)OSR(Z300_Conveyor[TMP_dConv].OSR_xRunMotor,Z300_Conveyor[TMP_dConv].OS_xRunMotor);